   "EMP IDB_stations_me{1}_partNumbers{5}" : WString[40] = PLC "EMP IDB".stations.me[1].partNumbers[5], 1 s
   "EMP IDB_stations_me{1}_partNumbers{6}" : WString[40] = PLC "EMP IDB".stations.me[1].partNumbers[6], 1 s
   "EMP IDB_stations_me{1}_partNumbers{7}" : WString[40] = PLC "EMP IDB".stations.me[1].partNumbers[7], 1 s
   "EMP IDB_stations_me{2}_partNumbers{0}" : WString[40] = PLC "EMP IDB".stations.me[2].partNumbers[0], 1 s
   "EMP IDB_stations_me{2}_partNumbers{1}" : WString[40] = PLC "EMP IDB".stations.me[2].partNumbers[1], 1 s
   "EMP IDB_stations_me{2}_partNumbers{2}" : WString[40] = PLC "EMP IDB".stations.me[2].partNumbers[2], 1 s
   "EMP IDB_stations_me{2}_partNumbers{3}" : WString[40] = PLC "EMP IDB".stations.me[2].partNumbers[3], 1 s
   "EMP IDB_stations_me{2}_partNumbers{4}" : WString[40] = PLC "EMP IDB".stations.me[2].partNumbers[4], 1 s
   "EMP IDB_stations_me{2}_partNumbers{5}" : WString[40] = PLC "EMP IDB".stations.me[2].partNumbers[5], 1 s
   "EMP IDB_stations_me{2}_partNumbers{6}" : WString[40] = PLC "EMP IDB".stations.me[2].partNumbers[6], 1 s
   "EMP IDB_stations_me{2}_partNumbers{7}" : WString[40] = PLC "EMP IDB".stations.me[2].partNumbers[7], 1 s
   "EMP IDB_stations_me{3}_partOrdered{0}" : Bool = PLC "EMP IDB".stations.me[3].partOrdered[0], 1 s
   "EMP IDB_stations_me{3}_partOrdered{1}" : Bool = PLC "EMP IDB".stations.me[3].partOrdered[1], 1 s
   "EMP IDB_stations_me{3}_partOrdered{2}" : Bool = PLC "EMP IDB".stations.me[3].partOrdered[2], 1 s
   "EMP IDB_stations_me{3}_partOrdered{3}" : Bool = PLC "EMP IDB".stations.me[3].partOrdered[3], 1 s
   "EMP IDB_stations_me{3}_partOrdered{4}" : Bool = PLC "EMP IDB".stations.me[3].partOrdered[4], 1 s
   "EMP IDB_stations_me{3}_partOrdered{5}" : Bool = PLC "EMP IDB".stations.me[3].partOrdered[5], 1 s
   "EMP IDB_stations_me{3}_partOrdered{6}" : Bool = PLC "EMP IDB".stations.me[3].partOrdered[6], 1 s
   "EMP IDB_stations_me{3}_partOrdered{7}" : Bool = PLC "EMP IDB".stations.me[3].partOrdered[7], 1 s
   "EMP IDB_stations_me{4}_partNumbers{0}" : WString[40] = PLC "EMP IDB".stations.me[4].partNumbers[0], 1 s
   "EMP IDB_stations_me{4}_partNumbers{1}" : WString[40] = PLC "EMP IDB".stations.me[4].partNumbers[1], 1 s
   "EMP IDB_stations_me{4}_partNumbers{2}" : WString[40] = PLC "EMP IDB".stations.me[4].partNumbers[2], 1 s
   "EMP IDB_stations_me{4}_partNumbers{3}" : WString[40] = PLC "EMP IDB".stations.me[4].partNumbers[3], 1 s
   "EMP IDB_stations_me{4}_partNumbers{4}" : WString[40] = PLC "EMP IDB".stations.me[4].partNumbers[4], 1 s
   "EMP IDB_stations_me{4}_partNumbers{5}" : WString[40] = PLC "EMP IDB".stations.me[4].partNumbers[5], 1 s
   "EMP IDB_stations_me{4}_partNumbers{6}" : WString[40] = PLC "EMP IDB".stations.me[4].partNumbers[6], 1 s
   "EMP IDB_stations_me{4}_partNumbers{7}" : WString[40] = PLC "EMP IDB".stations.me[4].partNumbers[7], 1 s
   "EMP IDB_stations_me{5}_partNumbers{0}" : WString[40] = PLC "EMP IDB".stations.me[5].partNumbers[0], 1 s
   "EMP IDB_stations_me{5}_partNumbers{1}" : WString[40] = PLC "EMP IDB".stations.me[5].partNumbers[1], 1 s
   "EMP IDB_stations_me{5}_partNumbers{2}" : WString[40] = PLC "EMP IDB".stations.me[5].partNumbers[2], 1 s
   "EMP IDB_stations_me{5}_partNumbers{3}" : WString[40] = PLC "EMP IDB".stations.me[5].partNumbers[3], 1 s
   "EMP IDB_stations_me{5}_partNumbers{4}" : WString[40] = PLC "EMP IDB".stations.me[5].partNumbers[4], 1 s
   "EMP IDB_stations_me{5}_partNumbers{5}" : WString[40] = PLC "EMP IDB".stations.me[5].partNumbers[5], 1 s
   "EMP IDB_stations_me{5}_partNumbers{6}" : WString[40] = PLC "EMP IDB".stations.me[5].partNumbers[6], 1 s
   "EMP IDB_stations_me{5}_partNumbers{7}" : WString[40] = PLC "EMP IDB".stations.me[5].partNumbers[7], 1 s
   "EMP IDB_stations_me{6}_partNumbers{0}" : WString[40] = PLC "EMP IDB".stations.me[6].partNumbers[0], 1 s
   "EMP IDB_stations_me{6}_partNumbers{1}" : WString[40] = PLC "EMP IDB".stations.me[6].partNumbers[1], 1 s
   "EMP IDB_stations_me{6}_partNumbers{2}" : WString[40] = PLC "EMP IDB".stations.me[6].partNumbers[2], 1 s
   "EMP IDB_stations_me{6}_partNumbers{3}" : WString[40] = PLC "EMP IDB".stations.me[6].partNumbers[3], 1 s
   "EMP IDB_stations_me{6}_partNumbers{4}" : WString[40] = PLC "EMP IDB".stations.me[6].partNumbers[4], 1 s
   "EMP IDB_stations_me{6}_partNumbers{5}" : WString[40] = PLC "EMP IDB".stations.me[6].partNumbers[5], 1 s
   "EMP IDB_stations_me{6}_partNumbers{6}" : WString[40] = PLC "EMP IDB".stations.me[6].partNumbers[6], 1 s
   "EMP IDB_stations_me{6}_partNumbers{7}" : WString[40] = PLC "EMP IDB".stations.me[6].partNumbers[7], 1 s
   "EMP IDB_stations_me{7}_partNumbers{0}" : WString[40] = PLC "EMP IDB".stations.me[7].partNumbers[0], 1 s
   "EMP IDB_stations_me{7}_partNumbers{1}" : WString[40] = PLC "EMP IDB".stations.me[7].partNumbers[1], 1 s
   "EMP IDB_stations_me{7}_partNumbers{2}" : WString[40] = PLC "EMP IDB".stations.me[7].partNumbers[2], 1 s
   "EMP IDB_stations_me{7}_partNumbers{3}" : WString[40] = PLC "EMP IDB".stations.me[7].partNumbers[3], 1 s
   "EMP IDB_stations_me{7}_partNumbers{4}" : WString[40] = PLC "EMP IDB".stations.me[7].partNumbers[4], 1 s
   "EMP IDB_stations_me{7}_partNumbers{5}" : WString[40] = PLC "EMP IDB".stations.me[7].partNumbers[5], 1 s
   "EMP IDB_stations_me{7}_partNumbers{6}" : WString[40] = PLC "EMP IDB".stations.me[7].partNumbers[6], 1 s
   "EMP IDB_stations_me{7}_partNumbers{7}" : WString[40] = PLC "EMP IDB".stations.me[7].partNumbers[7], 1 s
   "EMP IDB_stations_me{8}_partNumbers{0}" : WString[40] = PLC "EMP IDB".stations.me[8].partNumbers[0], 1 s
   "EMP IDB_stations_me{8}_partNumbers{1}" : WString[40] = PLC "EMP IDB".stations.me[8].partNumbers[1], 1 s
   "EMP IDB_stations_me{8}_partNumbers{2}" : WString[40] = PLC "EMP IDB".stations.me[8].partNumbers[2], 1 s
   "EMP IDB_stations_me{8}_partNumbers{3}" : WString[40] = PLC "EMP IDB".stations.me[8].partNumbers[3], 1 s
   "EMP IDB_stations_me{8}_partNumbers{4}" : WString[40] = PLC "EMP IDB".stations.me[8].partNumbers[4], 1 s
   "EMP IDB_stations_me{8}_partNumbers{5}" : WString[40] = PLC "EMP IDB".stations.me[8].partNumbers[5], 1 s
   "EMP IDB_stations_me{8}_partNumbers{6}" : WString[40] = PLC "EMP IDB".stations.me[8].partNumbers[6], 1 s
   "EMP IDB_stations_me{8}_partNumbers{7}" : WString[40] = PLC "EMP IDB".stations.me[8].partNumbers[7], 1 s
   "EMP IDB_stations_me{9}_partNumbers{0}" : WString[40] = PLC "EMP IDB".stations.me[9].partNumbers[0], 1 s
   "EMP IDB_stations_me{9}_partNumbers{1}" : WString[40] = PLC "EMP IDB".stations.me[9].partNumbers[1], 1 s
   "EMP IDB_stations_me{9}_partNumbers{2}" : WString[40] = PLC "EMP IDB".stations.me[9].partNumbers[2], 1 s
   "EMP IDB_stations_me{9}_partNumbers{3}" : WString[40] = PLC "EMP IDB".stations.me[9].partNumbers[3], 1 s
   "EMP IDB_stations_me{9}_partNumbers{4}" : WString[40] = PLC "EMP IDB".stations.me[9].partNumbers[4], 1 s
   "EMP IDB_stations_me{9}_partNumbers{5}" : WString[40] = PLC "EMP IDB".stations.me[9].partNumbers[5], 1 s
   "EMP IDB_stations_me{9}_partNumbers{6}" : WString[40] = PLC "EMP IDB".stations.me[9].partNumbers[6], 1 s
   "EMP IDB_stations_me{9}_partNumbers{7}" : WString[40] = PLC "EMP IDB".stations.me[9].partNumbers[7], 1 s
   "EMP IDB_stations_me{10}_partNumbers{0}" : WString[40] = PLC "EMP IDB".stations.me[10].partNumbers[0], 1 s
   "EMP IDB_stations_me{10}_partNumbers{1}" : WString[40] = PLC "EMP IDB".stations.me[10].partNumbers[1], 1 s
   "EMP IDB_stations_me{10}_partNumbers{2}" : WString[40] = PLC "EMP IDB".stations.me[10].partNumbers[2], 1 s
   "EMP IDB_stations_me{10}_partNumbers{3}" : WString[40] = PLC "EMP IDB".stations.me[10].partNumbers[3], 1 s
   "EMP IDB_stations_me{10}_partNumbers{4}" : WString[40] = PLC "EMP IDB".stations.me[10].partNumbers[4], 1 s
   "EMP IDB_stations_me{10}_partNumbers{5}" : WString[40] = PLC "EMP IDB".stations.me[10].partNumbers[5], 1 s
   "EMP IDB_stations_me{10}_partNumbers{6}" : WString[40] = PLC "EMP IDB".stations.me[10].partNumbers[6], 1 s
   "EMP IDB_stations_me{10}_partNumbers{7}" : WString[40] = PLC "EMP IDB".stations.me[10].partNumbers[7], 1 s
   "EMP IDB_stations_me{11}_partNumbers{0}" : WString[40] = PLC "EMP IDB".stations.me[11].partNumbers[0], 1 s
   "EMP IDB_stations_me{11}_partNumbers{1}" : WString[40] = PLC "EMP IDB".stations.me[11].partNumbers[1], 1 s
   "EMP IDB_stations_me{11}_partNumbers{2}" : WString[40] = PLC "EMP IDB".stations.me[11].partNumbers[2], 1 s
   "EMP IDB_stations_me{11}_partNumbers{3}" : WString[40] = PLC "EMP IDB".stations.me[11].partNumbers[3], 1 s
   "EMP IDB_stations_me{11}_partNumbers{4}" : WString[40] = PLC "EMP IDB".stations.me[11].partNumbers[4], 1 s
   "EMP IDB_stations_me{11}_partNumbers{5}" : WString[40] = PLC "EMP IDB".stations.me[11].partNumbers[5], 1 s
   "EMP IDB_stations_me{11}_partNumbers{6}" : WString[40] = PLC "EMP IDB".stations.me[11].partNumbers[6], 1 s
   "EMP IDB_stations_me{11}_partNumbers{7}" : WString[40] = PLC "EMP IDB".stations.me[11].partNumbers[7], 1 s
   "EMP IDB_stations_me{12}_partNumbers{0}" : WString[40] = PLC "EMP IDB".stations.me[12].partNumbers[0], 1 s
   "EMP IDB_stations_me{12}_partNumbers{1}" : WString[40] = PLC "EMP IDB".stations.me[12].partNumbers[1], 1 s
   "EMP IDB_stations_me{12}_partNumbers{2}" : WString[40] = PLC "EMP IDB".stations.me[12].partNumbers[2], 1 s
   "EMP IDB_stations_me{12}_partNumbers{3}" : WString[40] = PLC "EMP IDB".stations.me[12].partNumbers[3], 1 s
   "EMP IDB_stations_me{12}_partNumbers{4}" : WString[40] = PLC "EMP IDB".stations.me[12].partNumbers[4], 1 s
   "EMP IDB_stations_me{12}_partNumbers{5}" : WString[40] = PLC "EMP IDB".stations.me[12].partNumbers[5], 1 s
   "EMP IDB_stations_me{12}_partNumbers{6}" : WString[40] = PLC "EMP IDB".stations.me[12].partNumbers[6], 1 s
   "EMP IDB_stations_me{12}_partNumbers{7}" : WString[40] = PLC "EMP IDB".stations.me[12].partNumbers[7], 1 s
   "EMP IDB_stations_me{13}_partNumbers{0}" : WString[40] = PLC "EMP IDB".stations.me[13].partNumbers[0], 1 s
   "EMP IDB_stations_me{13}_partNumbers{1}" : WString[40] = PLC "EMP IDB".stations.me[13].partNumbers[1], 1 s
   "EMP IDB_stations_me{13}_partNumbers{2}" : WString[40] = PLC "EMP IDB".stations.me[13].partNumbers[2], 1 s
   "EMP IDB_stations_me{13}_partNumbers{3}" : WString[40] = PLC "EMP IDB".stations.me[13].partNumbers[3], 1 s
   "EMP IDB_stations_me{13}_partNumbers{4}" : WString[40] = PLC "EMP IDB".stations.me[13].partNumbers[4], 1 s
   "EMP IDB_stations_me{13}_partNumbers{5}" : WString[40] = PLC "EMP IDB".stations.me[13].partNumbers[5], 1 s
   "EMP IDB_stations_me{13}_partNumbers{6}" : WString[40] = PLC "EMP IDB".stations.me[13].partNumbers[6], 1 s
   "EMP IDB_stations_me{13}_partNumbers{7}" : WString[40] = PLC "EMP IDB".stations.me[13].partNumbers[7], 1 s
   "EMP IDB_stations_me{14}_partNumbers{0}" : WString[40] = PLC "EMP IDB".stations.me[14].partNumbers[0], 1 s
   "EMP IDB_stations_me{14}_partNumbers{1}" : WString[40] = PLC "EMP IDB".stations.me[14].partNumbers[1], 1 s
   "EMP IDB_stations_me{14}_partNumbers{2}" : WString[40] = PLC "EMP IDB".stations.me[14].partNumbers[2], 1 s
   "EMP IDB_stations_me{14}_partNumbers{3}" : WString[40] = PLC "EMP IDB".stations.me[14].partNumbers[3], 1 s
   "EMP IDB_stations_me{14}_partNumbers{4}" : WString[40] = PLC "EMP IDB".stations.me[14].partNumbers[4], 1 s
   "EMP IDB_stations_me{14}_partNumbers{5}" : WString[40] = PLC "EMP IDB".stations.me[14].partNumbers[5], 1 s
   "EMP IDB_stations_me{14}_partNumbers{6}" : WString[40] = PLC "EMP IDB".stations.me[14].partNumbers[6], 1 s
   "EMP IDB_stations_me{14}_partNumbers{7}" : WString[40] = PLC "EMP IDB".stations.me[14].partNumbers[7], 1 s
   "EMP IDB_stations_me{15}_partNumbers{0}" : WString[40] = PLC "EMP IDB".stations.me[15].partNumbers[0], 1 s
   "EMP IDB_stations_me{15}_partNumbers{1}" : WString[40] = PLC "EMP IDB".stations.me[15].partNumbers[1], 1 s
   "EMP IDB_stations_me{15}_partNumbers{2}" : WString[40] = PLC "EMP IDB".stations.me[15].partNumbers[2], 1 s
   "EMP IDB_stations_me{15}_partNumbers{3}" : WString[40] = PLC "EMP IDB".stations.me[15].partNumbers[3], 1 s
   "EMP IDB_stations_me{15}_partNumbers{4}" : WString[40] = PLC "EMP IDB".stations.me[15].partNumbers[4], 1 s
   "EMP IDB_stations_me{15}_partNumbers{5}" : WString[40] = PLC "EMP IDB".stations.me[15].partNumbers[5], 1 s
   "EMP IDB_stations_me{15}_partNumbers{6}" : WString[40] = PLC "EMP IDB".stations.me[15].partNumbers[6], 1 s
   "EMP IDB_stations_me{15}_partNumbers{7}" : WString[40] = PLC "EMP IDB".stations.me[15].partNumbers[7], 1 s
   "EMP IDB_stations_me{16}_partNumbers{0}" : WString[40] = PLC "EMP IDB".stations.me[16].partNumbers[0], 1 s
   "EMP IDB_stations_me{16}_partNumbers{1}" : WString[40] = PLC "EMP IDB".stations.me[16].partNumbers[1], 1 s
   "EMP IDB_stations_me{16}_partNumbers{2}" : WString[40] = PLC "EMP IDB".stations.me[16].partNumbers[2], 1 s
   "EMP IDB_stations_me{16}_partNumbers{3}" : WString[40] = PLC "EMP IDB".stations.me[16].partNumbers[3], 1 s
   "EMP IDB_stations_me{16}_partNumbers{4}" : WString[40] = PLC "EMP IDB".stations.me[16].partNumbers[4], 1 s
   "EMP IDB_stations_me{16}_partNumbers{5}" : WString[40] = PLC "EMP IDB".stations.me[16].partNumbers[5], 1 s
   "EMP IDB_stations_me{16}_partNumbers{6}" : WString[40] = PLC "EMP IDB".stations.me[16].partNumbers[6], 1 s
   "EMP IDB_stations_me{16}_partNumbers{7}" : WString[40] = PLC "EMP IDB".stations.me[16].partNumbers[7], 1 s
   "EMP IDB_stations_me{17}_partNumbers{0}" : WString[40] = PLC "EMP IDB".stations.me[17].partNumbers[0], 1 s
   "EMP IDB_stations_me{17}_partNumbers{1}" : WString[40] = PLC "EMP IDB".stations.me[17].partNumbers[1], 1 s
   "EMP IDB_stations_me{17}_partNumbers{2}" : WString[40] = PLC "EMP IDB".stations.me[17].partNumbers[2], 1 s
   "EMP IDB_stations_me{17}_partNumbers{3}" : WString[40] = PLC "EMP IDB".stations.me[17].partNumbers[3], 1 s
   "EMP IDB_stations_me{17}_partNumbers{4}" : WString[40] = PLC "EMP IDB".stations.me[17].partNumbers[4], 1 s
   "EMP IDB_stations_me{17}_partNumbers{5}" : WString[40] = PLC "EMP IDB".stations.me[17].partNumbers[5], 1 s
   "EMP IDB_stations_me{17}_partNumbers{6}" : WString[40] = PLC "EMP IDB".stations.me[17].partNumbers[6], 1 s
   "EMP IDB_stations_me{17}_partNumbers{7}" : WString[40] = PLC "EMP IDB".stations.me[17].partNumbers[7], 1 s
   "EMP IDB_stations_me{18}_partNumbers{0}" : WString[40] = PLC "EMP IDB".stations.me[18].partNumbers[0], 1 s
   "EMP IDB_stations_me{18}_partNumbers{1}" : WString[40] = PLC "EMP IDB".stations.me[18].partNumbers[1], 1 s
   "EMP IDB_stations_me{18}_partNumbers{2}" : WString[40] = PLC "EMP IDB".stations.me[18].partNumbers[2], 1 s
   "EMP IDB_stations_me{18}_partNumbers{3}" : WString[40] = PLC "EMP IDB".stations.me[18].partNumbers[3], 1 s
   "EMP IDB_stations_me{18}_partNumbers{4}" : WString[40] = PLC "EMP IDB".stations.me[18].partNumbers[4], 1 s
   "EMP IDB_stations_me{18}_partNumbers{5}" : WString[40] = PLC "EMP IDB".stations.me[18].partNumbers[5], 1 s
   "EMP IDB_stations_me{18}_partNumbers{6}" : WString[40] = PLC "EMP IDB".stations.me[18].partNumbers[6], 1 s
   "EMP IDB_stations_me{18}_partNumbers{7}" : WString[40] = PLC "EMP IDB".stations.me[18].partNumbers[7], 1 s
   "EMP IDB_stations_me{19}_partNumbers{0}" : WString[40] = PLC "EMP IDB".stations.me[19].partNumbers[0], 1 s
   "EMP IDB_stations_me{19}_partNumbers{1}" : WString[40] = PLC "EMP IDB".stations.me[19].partNumbers[1], 1 s
   "EMP IDB_stations_me{19}_partNumbers{2}" : WString[40] = PLC "EMP IDB".stations.me[19].partNumbers[2], 1 s
   "EMP IDB_stations_me{19}_partNumbers{3}" : WString[40] = PLC "EMP IDB".stations.me[19].partNumbers[3], 1 s
   "EMP IDB_stations_me{19}_partNumbers{4}" : WString[40] = PLC "EMP IDB".stations.me[19].partNumbers[4], 1 s
   "EMP IDB_stations_me{19}_partNumbers{5}" : WString[40] = PLC "EMP IDB".stations.me[19].partNumbers[5], 1 s
   "EMP IDB_stations_me{19}_partNumbers{6}" : WString[40] = PLC "EMP IDB".stations.me[19].partNumbers[6], 1 s
   "EMP IDB_stations_me{19}_partNumbers{7}" : WString[40] = PLC "EMP IDB".stations.me[19].partNumbers[7], 1 s
   "EMP IDB_stations_me{20}_partNumbers{0}" : WString[40] = PLC "EMP IDB".stations.me[20].partNumbers[0], 1 s
   "EMP IDB_stations_me{20}_partNumbers{1}" : WString[40] = PLC "EMP IDB".stations.me[20].partNumbers[1], 1 s
   "EMP IDB_stations_me{20}_partNumbers{2}" : WString[40] = PLC "EMP IDB".stations.me[20].partNumbers[2], 1 s
   "EMP IDB_stations_me{20}_partNumbers{3}" : WString[40] = PLC "EMP IDB".stations.me[20].partNumbers[3], 1 s
   "EMP IDB_stations_me{20}_partNumbers{4}" : WString[40] = PLC "EMP IDB".stations.me[20].partNumbers[4], 1 s
   "EMP IDB_stations_me{20}_partNumbers{5}" : WString[40] = PLC "EMP IDB".stations.me[20].partNumbers[5], 1 s
   "EMP IDB_stations_me{20}_partNumbers{6}" : WString[40] = PLC "EMP IDB".stations.me[20].partNumbers[6], 1 s
   "EMP IDB_stations_me{20}_partNumbers{7}" : WString[40] = PLC "EMP IDB".stations.me[20].partNumbers[7], 1 s
   "EMP IDB_stations_me{21}_partNumbers{0}" : WString[40] = PLC "EMP IDB".stations.me[21].partNumbers[0], 1 s
   "EMP IDB_stations_me{21}_partNumbers{1}" : WString[40] = PLC "EMP IDB".stations.me[21].partNumbers[1], 1 s
   "EMP IDB_stations_me{21}_partNumbers{2}" : WString[40] = PLC "EMP IDB".stations.me[21].partNumbers[2], 1 s
   "EMP IDB_stations_me{21}_partNumbers{3}" : WString[40] = PLC "EMP IDB".stations.me[21].partNumbers[3], 1 s
   "EMP IDB_stations_me{21}_partNumbers{4}" : WString[40] = PLC "EMP IDB".stations.me[21].partNumbers[4], 1 s
   "EMP IDB_stations_me{21}_partNumbers{5}" : WString[40] = PLC "EMP IDB".stations.me[21].partNumbers[5], 1 s
   "EMP IDB_stations_me{21}_partNumbers{6}" : WString[40] = PLC "EMP IDB".stations.me[21].partNumbers[6], 1 s
   "EMP IDB_stations_me{21}_partNumbers{7}" : WString[40] = PLC "EMP IDB".stations.me[21].partNumbers[7], 1 s
   "EMP IDB_stations_me{22}_partNumbers{0}" : WString[40] = PLC "EMP IDB".stations.me[22].partNumbers[0], 1 s
   "EMP IDB_stations_me{22}_partNumbers{1}" : WString[40] = PLC "EMP IDB".stations.me[22].partNumbers[1], 1 s
   "EMP IDB_stations_me{22}_partNumbers{2}" : WString[40] = PLC "EMP IDB".stations.me[22].partNumbers[2], 1 s
   "EMP IDB_stations_me{22}_partNumbers{3}" : WString[40] = PLC "EMP IDB".stations.me[22].partNumbers[3], 1 s
   "EMP IDB_stations_me{22}_partNumbers{4}" : WString[40] = PLC "EMP IDB".stations.me[22].partNumbers[4], 1 s
   "EMP IDB_stations_me{22}_partNumbers{5}" : WString[40] = PLC "EMP IDB".stations.me[22].partNumbers[5], 1 s
   "EMP IDB_stations_me{22}_partNumbers{6}" : WString[40] = PLC "EMP IDB".stations.me[22].partNumbers[6], 1 s
   "EMP IDB_stations_me{22}_partNumbers{7}" : WString[40] = PLC "EMP IDB".stations.me[22].partNumbers[7], 1 s
   "EMP IDB_stations_me{23}_partNumbers{0}" : WString[40] = PLC "EMP IDB".stations.me[23].partNumbers[0], 1 s
   "EMP IDB_stations_me{23}_partNumbers{1}" : WString[40] = PLC "EMP IDB".stations.me[23].partNumbers[1], 1 s
   "EMP IDB_stations_me{23}_partNumbers{2}" : WString[40] = PLC "EMP IDB".stations.me[23].partNumbers[2], 1 s
   "EMP IDB_stations_me{23}_partNumbers{3}" : WString[40] = PLC "EMP IDB".stations.me[23].partNumbers[3], 1 s
   "EMP IDB_stations_me{23}_partNumbers{4}" : WString[40] = PLC "EMP IDB".stations.me[23].partNumbers[4], 1 s
   "EMP IDB_stations_me{23}_partNumbers{5}" : WString[40] = PLC "EMP IDB".stations.me[23].partNumbers[5], 1 s
   "EMP IDB_stations_me{23}_partNumbers{6}" : WString[40] = PLC "EMP IDB".stations.me[23].partNumbers[6], 1 s
   "EMP IDB_stations_me{23}_partNumbers{7}" : WString[40] = PLC "EMP IDB".stations.me[23].partNumbers[7], 1 s
   "EMP IDB_stations_me{3}_partNumbers{0}" : WString[40] = PLC "EMP IDB".stations.me[3].partNumbers[0], 1 s
   "EMP IDB_stations_me{3}_partNumbers{1}" : WString[40] = PLC "EMP IDB".stations.me[3].partNumbers[1], 1 s
   "EMP IDB_stations_me{3}_partNumbers{2}" : WString[40] = PLC "EMP IDB".stations.me[3].partNumbers[2], 1 s
   "EMP IDB_stations_me{3}_partNumbers{3}" : WString[40] = PLC "EMP IDB".stations.me[3].partNumbers[3], 1 s
   "EMP IDB_stations_me{3}_partNumbers{4}" : WString[40] = PLC "EMP IDB".stations.me[3].partNumbers[4], 1 s
   "EMP IDB_stations_me{3}_partNumbers{5}" : WString[40] = PLC "EMP IDB".stations.me[3].partNumbers[5], 1 s
   "EMP IDB_stations_me{3}_partNumbers{6}" : WString[40] = PLC "EMP IDB".stations.me[3].partNumbers[6], 1 s
   "EMP IDB_stations_me{3}_partNumbers{7}" : WString[40] = PLC "EMP IDB".stations.me[3].partNumbers[7], 1 s

text list "Station Selection Single": 0 'Select a Station to View'; 1 'Assignments'

recipe "VOLVO 16 01": Button 0 <- "EMP IDB_stations_me{0}_partNumbers{0}", Button 1 <- "EMP IDB_stations_me{0}_partNumbers{1}", Button 2 <- "EMP IDB_stations_me{0}_partNumbers{2}", Button 3 <- "EMP IDB_stations_me{0}_partNumbers{3}", Button 4 <- "EMP IDB_stations_me{0}_partNumbers{4}", Button 5 <- "EMP IDB_stations_me{0}_partNumbers{5}", Button 6 <- "EMP IDB_stations_me{0}_partNumbers{6}", Button 7 <- "EMP IDB_stations_me{0}_partNumbers{7}"

recipe "VOLVO 16 02": Button 0 <- "EMP IDB_stations_me{1}_partNumbers{0}", Button 1 <- "EMP IDB_stations_me{1}_partNumbers{1}", Button 2 <- "EMP IDB_stations_me{1}_partNumbers{2}", Button 3 <- "EMP IDB_stations_me{1}_partNumbers{3}", Button 4 <- "EMP IDB_stations_me{1}_partNumbers{4}", Button 5 <- "EMP IDB_stations_me{1}_partNumbers{5}", Button 6 <- "EMP IDB_stations_me{1}_partNumbers{6}", Button 7 <- "EMP IDB_stations_me{1}_partNumbers{7}"

recipe "VOLVO 16 03": Button 0 <- "EMP IDB_stations_me{2}_partNumbers{0}", Button 1 <- "EMP IDB_stations_me{2}_partNumbers{1}", Button 2 <- "EMP IDB_stations_me{2}_partNumbers{2}", Button 3 <- "EMP IDB_stations_me{2}_partNumbers{3}", Button 4 <- "EMP IDB_stations_me{2}_partNumbers{4}", Button 5 <- "EMP IDB_stations_me{2}_partNumbers{5}", Button 6 <- "EMP IDB_stations_me{2}_partNumbers{6}", Button 7 <- "EMP IDB_stations_me{2}_partNumbers{7}"

recipe "VOLVO 16 04": Button 0 <- "EMP IDB_stations_me{3}_partNumbers{0}", Button 1 <- "EMP IDB_stations_me{3}_partNumbers{1}", Button 2 <- "EMP IDB_stations_me{3}_partNumbers{2}", Button 3 <- "EMP IDB_stations_me{3}_partNumbers{3}", Button 4 <- "EMP IDB_stations_me{3}_partNumbers{4}", Button 5 <- "EMP IDB_stations_me{3}_partNumbers{5}", Button 6 <- "EMP IDB_stations_me{3}_partNumbers{6}", Button 7 <- "EMP IDB_stations_me{3}_partNumbers{7}"

recipe "VOLVO 16 05": Button 0 <- "EMP IDB_stations_me{4}_partNumbers{0}", Button 1 <- "EMP IDB_stations_me{4}_partNumbers{1}", Button 2 <- "EMP IDB_stations_me{4}_partNumbers{2}", Button 3 <- "EMP IDB_stations_me{4}_partNumbers{3}", Button 4 <- "EMP IDB_stations_me{4}_partNumbers{4}", Button 5 <- "EMP IDB_stations_me{4}_partNumbers{5}", Button 6 <- "EMP IDB_stations_me{4}_partNumbers{6}", Button 7 <- "EMP IDB_stations_me{4}_partNumbers{7}"

recipe "VOLVO 16 06": Button 0 <- "EMP IDB_stations_me{5}_partNumbers{0}", Button 1 <- "EMP IDB_stations_me{5}_partNumbers{1}", Button 2 <- "EMP IDB_stations_me{5}_partNumbers{2}", Button 3 <- "EMP IDB_stations_me{5}_partNumbers{3}", Button 4 <- "EMP IDB_stations_me{5}_partNumbers{4}", Button 5 <- "EMP IDB_stations_me{5}_partNumbers{5}", Button 6 <- "EMP IDB_stations_me{5}_partNumbers{6}", Button 7 <- "EMP IDB_stations_me{5}_partNumbers{7}"

recipe "VOLVO 16 07": Button 0 <- "EMP IDB_stations_me{6}_partNumbers{0}", Button 1 <- "EMP IDB_stations_me{6}_partNumbers{1}", Button 2 <- "EMP IDB_stations_me{6}_partNumbers{2}", Button 3 <- "EMP IDB_stations_me{6}_partNumbers{3}", Button 4 <- "EMP IDB_stations_me{6}_partNumbers{4}", Button 5 <- "EMP IDB_stations_me{6}_partNumbers{5}", Button 6 <- "EMP IDB_stations_me{6}_partNumbers{6}", Button 7 <- "EMP IDB_stations_me{6}_partNumbers{7}"

recipe "VOLVO 16 08": Button 0 <- "EMP IDB_stations_me{7}_partNumbers{0}", Button 1 <- "EMP IDB_stations_me{7}_partNumbers{1}", Button 2 <- "EMP IDB_stations_me{7}_partNumbers{2}", Button 3 <- "EMP IDB_stations_me{7}_partNumbers{3}", Button 4 <- "EMP IDB_stations_me{7}_partNumbers{4}", Button 5 <- "EMP IDB_stations_me{7}_partNumbers{5}", Button 6 <- "EMP IDB_stations_me{7}_partNumbers{6}", Button 7 <- "EMP IDB_stations_me{7}_partNumbers{7}"

recipe "VOLVO 16 09": Button 0 <- "EMP IDB_stations_me{8}_partNumbers{0}", Button 1 <- "EMP IDB_stations_me{8}_partNumbers{1}", Button 2 <- "EMP IDB_stations_me{8}_partNumbers{2}", Button 3 <- "EMP IDB_stations_me{8}_partNumbers{3}", Button 4 <- "EMP IDB_stations_me{8}_partNumbers{4}", Button 5 <- "EMP IDB_stations_me{8}_partNumbers{5}", Button 6 <- "EMP IDB_stations_me{8}_partNumbers{6}", Button 7 <- "EMP IDB_stations_me{8}_partNumbers{7}"

recipe "VOLVO 16 10": Button 0 <- "EMP IDB_stations_me{9}_partNumbers{0}", Button 1 <- "EMP IDB_stations_me{9}_partNumbers{1}", Button 2 <- "EMP IDB_stations_me{9}_partNumbers{2}", Button 3 <- "EMP IDB_stations_me{9}_partNumbers{3}", Button 4 <- "EMP IDB_stations_me{9}_partNumbers{4}", Button 5 <- "EMP IDB_stations_me{9}_partNumbers{5}", Button 6 <- "EMP IDB_stations_me{9}_partNumbers{6}", Button 7 <- "EMP IDB_stations_me{9}_partNumbers{7}"

recipe "VOLVO 16 11": Button 0 <- "EMP IDB_stations_me{10}_partNumbers{0}", Button 1 <- "EMP IDB_stations_me{10}_partNumbers{1}", Button 2 <- "EMP IDB_stations_me{10}_partNumbers{2}", Button 3 <- "EMP IDB_stations_me{10}_partNumbers{3}", Button 4 <- "EMP IDB_stations_me{10}_partNumbers{4}", Button 5 <- "EMP IDB_stations_me{10}_partNumbers{5}", Button 6 <- "EMP IDB_stations_me{10}_partNumbers{6}", Button 7 <- "EMP IDB_stations_me{10}_partNumbers{7}"

recipe "CHM 01": Button 0 <- "EMP IDB_stations_me{11}_partNumbers{0}", Button 1 <- "EMP IDB_stations_me{11}_partNumbers{1}", Button 2 <- "EMP IDB_stations_me{11}_partNumbers{2}", Button 3 <- "EMP IDB_stations_me{11}_partNumbers{3}", Button 4 <- "EMP IDB_stations_me{11}_partNumbers{4}", Button 5 <- "EMP IDB_stations_me{11}_partNumbers{5}", Button 6 <- "EMP IDB_stations_me{11}_partNumbers{6}", Button 7 <- "EMP IDB_stations_me{11}_partNumbers{7}"

recipe "CHM 02": Button 0 <- "EMP IDB_stations_me{12}_partNumbers{0}", Button 1 <- "EMP IDB_stations_me{12}_partNumbers{1}", Button 2 <- "EMP IDB_stations_me{12}_partNumbers{2}", Button 3 <- "EMP IDB_stations_me{12}_partNumbers{3}", Button 4 <- "EMP IDB_stations_me{12}_partNumbers{4}", Button 5 <- "EMP IDB_stations_me{12}_partNumbers{5}", Button 6 <- "EMP IDB_stations_me{12}_partNumbers{6}", Button 7 <- "EMP IDB_stations_me{12}_partNumbers{7}"

recipe "CHM 03": Button 0 <- "EMP IDB_stations_me{13}_partNumbers{0}", Button 1 <- "EMP IDB_stations_me{13}_partNumbers{1}", Button 2 <- "EMP IDB_stations_me{13}_partNumbers{2}", Button 3 <- "EMP IDB_stations_me{13}_partNumbers{3}", Button 4 <- "EMP IDB_stations_me{13}_partNumbers{4}", Button 5 <- "EMP IDB_stations_me{13}_partNumbers{5}", Button 6 <- "EMP IDB_stations_me{13}_partNumbers{6}", Button 7 <- "EMP IDB_stations_me{13}_partNumbers{7}"

recipe "CHM 04": Button 0 <- "EMP IDB_stations_me{14}_partNumbers{0}", Button 1 <- "EMP IDB_stations_me{14}_partNumbers{1}", Button 2 <- "EMP IDB_stations_me{14}_partNumbers{2}", Button 3 <- "EMP IDB_stations_me{14}_partNumbers{3}", Button 4 <- "EMP IDB_stations_me{14}_partNumbers{4}", Button 5 <- "EMP IDB_stations_me{14}_partNumbers{5}", Button 6 <- "EMP IDB_stations_me{14}_partNumbers{6}", Button 7 <- "EMP IDB_stations_me{14}_partNumbers{7}"

recipe "CHM 05": Button 0 <- "EMP IDB_stations_me{15}_partNumbers{0}", Button 1 <- "EMP IDB_stations_me{15}_partNumbers{1}", Button 2 <- "EMP IDB_stations_me{15}_partNumbers{2}", Button 3 <- "EMP IDB_stations_me{15}_partNumbers{3}", Button 4 <- "EMP IDB_stations_me{15}_partNumbers{4}", Button 5 <- "EMP IDB_stations_me{15}_partNumbers{5}", Button 6 <- "EMP IDB_stations_me{15}_partNumbers{6}", Button 7 <- "EMP IDB_stations_me{15}_partNumbers{7}"

recipe "CDO 01": Button 0 <- "EMP IDB_stations_me{16}_partNumbers{0}", Button 1 <- "EMP IDB_stations_me{16}_partNumbers{1}", Button 2 <- "EMP IDB_stations_me{16}_partNumbers{2}", Button 3 <- "EMP IDB_stations_me{16}_partNumbers{3}", Button 4 <- "EMP IDB_stations_me{16}_partNumbers{4}", Button 5 <- "EMP IDB_stations_me{16}_partNumbers{5}", Button 6 <- "EMP IDB_stations_me{16}_partNumbers{6}", Button 7 <- "EMP IDB_stations_me{16}_partNumbers{7}"

recipe "CDO 02": Button 0 <- "EMP IDB_stations_me{17}_partNumbers{0}", Button 1 <- "EMP IDB_stations_me{17}_partNumbers{1}", Button 2 <- "EMP IDB_stations_me{17}_partNumbers{2}", Button 3 <- "EMP IDB_stations_me{17}_partNumbers{3}", Button 4 <- "EMP IDB_stations_me{17}_partNumbers{4}", Button 5 <- "EMP IDB_stations_me{17}_partNumbers{5}", Button 6 <- "EMP IDB_stations_me{17}_partNumbers{6}", Button 7 <- "EMP IDB_stations_me{17}_partNumbers{7}"

recipe "CDO 03": Button 0 <- "EMP IDB_stations_me{18}_partNumbers{0}", Button 1 <- "EMP IDB_stations_me{18}_partNumbers{1}", Button 2 <- "EMP IDB_stations_me{18}_partNumbers{2}", Button 3 <- "EMP IDB_stations_me{18}_partNumbers{3}", Button 4 <- "EMP IDB_stations_me{18}_partNumbers{4}", Button 5 <- "EMP IDB_stations_me{18}_partNumbers{5}", Button 6 <- "EMP IDB_stations_me{18}_partNumbers{6}", Button 7 <- "EMP IDB_stations_me{18}_partNumbers{7}"

recipe "BFL 01": Button 0 <- "EMP IDB_stations_me{19}_partNumbers{0}", Button 1 <- "EMP IDB_stations_me{19}_partNumbers{1}", Button 2 <- "EMP IDB_stations_me{19}_partNumbers{2}", Button 3 <- "EMP IDB_stations_me{19}_partNumbers{3}", Button 4 <- "EMP IDB_stations_me{19}_partNumbers{4}", Button 5 <- "EMP IDB_stations_me{19}_partNumbers{5}", Button 6 <- "EMP IDB_stations_me{19}_partNumbers{6}", Button 7 <- "EMP IDB_stations_me{19}_partNumbers{7}"

recipe "BFL 02": Button 0 <- "EMP IDB_stations_me{20}_partNumbers{0}", Button 1 <- "EMP IDB_stations_me{20}_partNumbers{1}", Button 2 <- "EMP IDB_stations_me{20}_partNumbers{2}", Button 3 <- "EMP IDB_stations_me{20}_partNumbers{3}", Button 4 <- "EMP IDB_stations_me{20}_partNumbers{4}", Button 5 <- "EMP IDB_stations_me{20}_partNumbers{5}", Button 6 <- "EMP IDB_stations_me{20}_partNumbers{6}", Button 7 <- "EMP IDB_stations_me{20}_partNumbers{7}"

recipe "BFL 03": Button 0 <- "EMP IDB_stations_me{21}_partNumbers{0}", Button 1 <- "EMP IDB_stations_me{21}_partNumbers{1}", Button 2 <- "EMP IDB_stations_me{21}_partNumbers{2}", Button 3 <- "EMP IDB_stations_me{21}_partNumbers{3}", Button 4 <- "EMP IDB_stations_me{21}_partNumbers{4}", Button 5 <- "EMP IDB_stations_me{21}_partNumbers{5}", Button 6 <- "EMP IDB_stations_me{21}_partNumbers{6}", Button 7 <- "EMP IDB_stations_me{21}_partNumbers{7}"

recipe "LGS 01": Button 0 <- "EMP IDB_stations_me{22}_partNumbers{0}", Button 1 <- "EMP IDB_stations_me{22}_partNumbers{1}", Button 2 <- "EMP IDB_stations_me{22}_partNumbers{2}", Button 3 <- "EMP IDB_stations_me{22}_partNumbers{3}", Button 4 <- "EMP IDB_stations_me{22}_partNumbers{4}", Button 5 <- "EMP IDB_stations_me{22}_partNumbers{5}", Button 6 <- "EMP IDB_stations_me{22}_partNumbers{6}", Button 7 <- "EMP IDB_stations_me{22}_partNumbers{7}"

recipe "LGS 02": Button 0 <- "EMP IDB_stations_me{23}_partNumbers{0}", Button 1 <- "EMP IDB_stations_me{23}_partNumbers{1}", Button 2 <- "EMP IDB_stations_me{23}_partNumbers{2}", Button 3 <- "EMP IDB_stations_me{23}_partNumbers{3}", Button 4 <- "EMP IDB_stations_me{23}_partNumbers{4}", Button 5 <- "EMP IDB_stations_me{23}_partNumbers{5}", Button 6 <- "EMP IDB_stations_me{23}_partNumbers{6}", Button 7 <- "EMP IDB_stations_me{23}_partNumbers{7}"

screen "1 PART CALL" 1366x768
   on GenerateScreen: SetTag("HMI_screenNumber", 1)
   Rectangle "Settings Tab Background" at 682,0 size 684x68
      Appearance <- "HMI_screenNumber"
   Rectangle "Part Call Tab Background" at 0,0 size 685x68
      Appearance <- "HMI_screenNumber"
   Rectangle "Settings Tab Border Hide" at 685,61 size 678x20
      Visibility <- "HMI_screenNumber"
   Rectangle "Part Call Tab Border Hide" at 3,61 size 679x20
      Visibility <- "HMI_screenNumber"
   Button "Settings Screen" at 683,0 size 683x68; TextOff 'SETTINGS'; Authorization "User administration"
      on Release: ActivateScreen("2 SETTINGS", 0)
   Button "Part Call Screen" at 0,0 size 683x68; TextOff 'PART CALL'
      on Release: ActivateScreen("1 PART CALL", 0)
   TextField "Header Line" at 32,112 size 216x53; Text 'LINE'
   TextField "Header Drop Zone" at 238,112 size 236x53; Text 'DROP ZONE'
   TextField "Header Part Number" at 474,112 size 648x53; Text 'PART NUMBER'
   TextField "Header Time" at 1112,112 size 222x53; Text 'TIME'
   ScreenModuleView "TableRow00" at 27,170 size 1312x52; ScreenModuleType ""
      Guid_{11997190-27688} <- "HMI_partCall_row{0}"
      on Guid_{11997190-83214}: ActivateScreen("3 BARCODE", 0)
   ScreenModuleView "TableRow01" at 27,222 size 1312x52; ScreenModuleType ""
      Guid_{11997190-27688} <- "HMI_partCall_row{1}"
      on Guid_{11997190-83214}: ActivateScreen("3 BARCODE", 0)
   ScreenModuleView "TableRow02" at 27,274 size 1312x52; ScreenModuleType ""
      Guid_{11997190-27688} <- "HMI_partCall_row{2}"
      on Guid_{11997190-83214}: ActivateScreen("3 BARCODE", 0)
   ScreenModuleView "TableRow03" at 27,326 size 1312x52; ScreenModuleType ""
      Guid_{11997190-27688} <- "HMI_partCall_row{3}"
      on Guid_{11997190-83214}: ActivateScreen("3 BARCODE", 0)
   ScreenModuleView "TableRow04" at 27,378 size 1312x52; ScreenModuleType ""
      Guid_{11997190-27688} <- "HMI_partCall_row{4}"
      on Guid_{11997190-83214}: ActivateScreen("3 BARCODE", 0)
   ScreenModuleView "TableRow05" at 27,430 size 1312x52; ScreenModuleType ""
      Guid_{11997190-27688} <- "HMI_partCall_row{5}"
      on Guid_{11997190-83214}: ActivateScreen("3 BARCODE", 0)
   ScreenModuleView "TableRow06" at 27,482 size 1312x52; ScreenModuleType ""
      Guid_{11997190-27688} <- "HMI_partCall_row{6}"
      on Guid_{11997190-83214}: ActivateScreen("3 BARCODE", 0)
   ScreenModuleView "TableRow07" at 27,534 size 1312x52; ScreenModuleType ""
      Guid_{11997190-27688} <- "HMI_partCall_row{7}"
      on Guid_{11997190-83214}: ActivateScreen("3 BARCODE", 0)
   ScreenModuleView "TableRow08" at 27,586 size 1312x52; ScreenModuleType ""
      Guid_{11997190-27688} <- "HMI_partCall_row{8}"
      on Guid_{11997190-83214}: ActivateScreen("3 BARCODE", 0)
   ScreenModuleView "TableRow09" at 27,638 size 1312x52; ScreenModuleType ""
      Guid_{11997190-27688} <- "HMI_partCall_row{9}"
      on Guid_{11997190-83214}: ActivateScreen("3 BARCODE", 0)
   ScreenModuleView "TableRow10" at 27,690 size 1312x52; ScreenModuleType ""
      Guid_{11997190-27688} <- "HMI_partCall_row{10}"
      on Guid_{11997190-83214}: ActivateScreen("3 BARCODE", 0)

screen "2 SETTINGS" 1366x768
   on GenerateScreen: SetTag("HMI_screenNumber", 2)
   Rectangle "Part Call Nave Panel" at 0,0 size 455x68
      Appearance <- "HMI_screenNumber"
   Rectangle "Settings Nav Panel" at 452,0 size 462x68
      Appearance <- "HMI_screenNumber"
   Rectangle "Network Health Nav Panel" at 911,0 size 455x68
      Appearance <- "HMI_screenNumber"
   Rectangle "Part Call Border Hide" at 3,60 size 449x20
      Visibility <- "HMI_screenNumber"
   Rectangle "Settings Border Hide" at 455,60 size 456x20
      Visibility <- "HMI_screenNumber"
   Rectangle "Network Health Border Hide" at 914,60 size 449x20
      Visibility <- "HMI_screenNumber"
   Button "Part Call Screen" at 0,0 size 455x68; TextOff 'PART CALL'
      on Release: ActivateScreen("1 PART CALL", 0)
   Button "Settings Screen" at 455,0 size 460x68; TextOff 'SETTINGS'
      on Release: ActivateScreen("2 SETTINGS", 0)
   Button "Network Health Screen" at 914,0 size 452x68; TextOff 'NW HEALTH'
      on Release: ActivateScreen("4 NETWORK HEALTH", 0)
   Rectangle "Station Assignment Table BG Full" at 793,120 size 533x630
      Visibility <- "HMI_settings_stations_selCount"
   TextField "Current Station Single" at 803,130 size 513x45; Text 'Text'
      Visibility <- "HMI_settings_stations_selCount"
   TextField "Hide Line and Drop Zone Multi" at 803,181 size 513x40; Text 'select single station for Line and Drop Zone'
      Visibility <- "HMI_settings_stations_selCount"
   GraphicView "KP8 Image" at 496,327 size 275x412; Picture "kp8 image"
   Rectangle "Station Assignment Table BG Mini" at 793,120 size 533x65
      Visibility <- "HMI_settings_stations_selCount"
   ScreenModuleView "PB: Set PN" at 50,130 size 414x45; Guid_{11997190-63616} 'Assign Part Number'; ScreenModuleType ""
      Guid_{11997190-63605} <- "HMI_settings_partNumber_assign"
   ScreenModuleView "PN IO Field" at 50,180 size 414x50; ScreenModuleType ""
      Guid_{11997190-63113} <- "HMI_settings_partNumber_ioField"
   ScreenModuleView "PB: Set Allotted" at 494,130 size 137x45; Guid_{11997190-63616} 'Allotted'; ScreenModuleType ""
      Guid_{11997190-63605} <- "HMI_settings_alotted_assign"
   ScreenModuleView "PB: Set Critical" at 636,130 size 137x45; Guid_{11997190-63616} 'Crititcal'; ScreenModuleType ""
      Guid_{11997190-63605} <- "HMI_settings_critical_assign"
   ScreenModuleView "Alotted Time IO Field" at 494,180 size 137x50; ScreenModuleType ""
      Guid_{11997190-63269} <- "HMI_settings_alotted_ioField"
   ScreenModuleView "Critical Time IO Field" at 636,180 size 137x50; ScreenModuleType ""
      Guid_{11997190-63269} <- "HMI_settings_critical_ioField"
   ScreenModuleView "PB: Select KP8 Buttons" at 493,270 size 284x45; Guid_{11997190-63616} 'Select Buttons'; ScreenModuleType ""
      Guid_{11997190-63605} <- "HMI_settings_kp8_selectButtons"
   ScreenModuleView "KP8 00: RESET" at 641,614 size 68x66; ScreenModuleType ""
      Guid_{11997190-57808} <- "HMI_settings_kp8_buttons{0}"
   ScreenModuleView "KP8 01" at 641,535 size 68x66; ScreenModuleType ""
      Guid_{11997190-57808} <- "HMI_settings_kp8_buttons{1}"
   ScreenModuleView "KP8 02" at 641,459 size 68x66; ScreenModuleType ""
      Guid_{11997190-57808} <- "HMI_settings_kp8_buttons{2}"
   ScreenModuleView "KP8 03" at 641,383 size 68x66; ScreenModuleType ""
      Guid_{11997190-57808} <- "HMI_settings_kp8_buttons{3}"
   ScreenModuleView "KP8 04: STOP RUNTIME" at 557,614 size 68x66; ScreenModuleType ""
      on Guid_{11997190-59171}: StopRuntime(0)
      Guid_{11997190-57808} <- "HMI_settings_kp8_buttons{4}"
   ScreenModuleView "KP8 05" at 557,535 size 68x66; ScreenModuleType ""
      Guid_{11997190-57808} <- "HMI_settings_kp8_buttons{5}"
   ScreenModuleView "KP8 06" at 557,459 size 68x66; ScreenModuleType ""
      Guid_{11997190-57808} <- "HMI_settings_kp8_buttons{6}"
   ScreenModuleView "KP8 07" at 557,383 size 68x66; ScreenModuleType ""
      Guid_{11997190-57808} <- "HMI_settings_kp8_buttons{7}"
   ScreenModuleView "PB: Previous Group" at 50,270 size 65x45; Guid_{11997190-63799} "Up"; ScreenModuleType ""
      Guid_{11997190-63779} <- "HMI_settings_stations_prevGroup"
   ScreenModuleView "PB: Select All Stations" at 120,270 size 274x45; Guid_{11997190-63616} 'Select Stations'; ScreenModuleType ""
      Guid_{11997190-63605} <- "HMI_settings_stations_selectAll"
   ScreenModuleView "PB: Next Group" at 399,270 size 65x45; Guid_{11997190-63799} "Down"; ScreenModuleType ""
      Guid_{11997190-63779} <- "HMI_settings_stations_nextGroup"
   ScreenModuleView "Station 00 Select" at 50,320 size 205x65; ScreenModuleType ""
      Guid_{11997190-57808} <- "HMI_settings_stations_selectBtns{0}"
   ScreenModuleView "Station 01 Select" at 260,320 size 205x65; ScreenModuleType ""
      Guid_{11997190-57808} <- "HMI_settings_stations_selectBtns{1}"
   ScreenModuleView "Station 02 Select" at 50,391 size 205x65; ScreenModuleType ""
      Guid_{11997190-57808} <- "HMI_settings_stations_selectBtns{2}"
   ScreenModuleView "Station 03 Select" at 260,391 size 205x65; ScreenModuleType ""
      Guid_{11997190-57808} <- "HMI_settings_stations_selectBtns{3}"
   ScreenModuleView "Station 04 Select" at 50,462 size 205x65; ScreenModuleType ""
      Guid_{11997190-57808} <- "HMI_settings_stations_selectBtns{4}"
   ScreenModuleView "Station 05 Select" at 260,462 size 205x65; ScreenModuleType ""
      Guid_{11997190-57808} <- "HMI_settings_stations_selectBtns{5}"
   ScreenModuleView "Station 06 Select" at 50,533 size 205x65; ScreenModuleType ""
      Guid_{11997190-57808} <- "HMI_settings_stations_selectBtns{6}"
   ScreenModuleView "Station 07 Select" at 260,533 size 205x65; ScreenModuleType ""
      Guid_{11997190-57808} <- "HMI_settings_stations_selectBtns{7}"
   ScreenModuleView "Station 08 Select" at 50,604 size 205x65; ScreenModuleType ""
      Guid_{11997190-57808} <- "HMI_settings_stations_selectBtns{8}"
   ScreenModuleView "Station 09 Select" at 260,604 size 205x65; ScreenModuleType ""
      Guid_{11997190-57808} <- "HMI_settings_stations_selectBtns{9}"
   ScreenModuleView "Station 10 Select" at 50,675 size 205x65; ScreenModuleType ""
      Guid_{11997190-57808} <- "HMI_settings_stations_selectBtns{10}"
   ScreenModuleView "Station 11 Select" at 260,675 size 205x65; ScreenModuleType ""
      Guid_{11997190-57808} <- "HMI_settings_stations_selectBtns{11}"
   ScreenModuleView "Line Label" at 803,181 size 267x40; ScreenModuleType ""
      Guid_{11997190-64598} <- "HMI_settings_viewingStation_lineData"
   ScreenModuleView "Drop Zone Label" at 1076,181 size 240x40; ScreenModuleType ""
      Guid_{11997190-64802} <- "HMI_settings_viewingStation_dzData"
   ScreenModuleView "PB: Previous Station" at 803,130 size 65x45; Guid_{11997190-63799} "Left"; ScreenModuleType ""
      Guid_{11997190-63779} <- "HMI_settings_viewingStation_previous"
   TextField "Current Station Multi" at 873,130 size 373x45; Text 'Assignments'
      Visibility <- "HMI_settings_stations_selCount"
   ScreenModuleView "PB: Next Station" at 1251,130 size 65x45; Guid_{11997190-63799} "Right"; ScreenModuleType ""
      Guid_{11997190-63779} <- "HMI_settings_viewingStation_next"
   TextField "Button Column Header" at 803,226 size 75x40; Text 'Btn'
      Visibility <- "HMI_settings_stations_selCount"
   TextField "Timer Column Header" at 872,226 size 128x40; Text 'Times'
      Visibility <- "HMI_settings_stations_selCount"
   TextField "Part Number Column Header" at 993,226 size 323x40; Text 'Part Number'
      Visibility <- "HMI_settings_stations_selCount"
   ScreenModuleView "Button 00 Details" at 803,271 size 513x74; ScreenModuleType ""
      Guid_{11997190-60358} <- "HMI_settings_viewingStation_btns{0}"
   ScreenModuleView "Button 01 Details" at 803,350 size 513x74; ScreenModuleType ""
      Guid_{11997190-60358} <- "HMI_settings_viewingStation_btns{1}"
   ScreenModuleView "Button 02 Details" at 803,429 size 513x74; ScreenModuleType ""
      Guid_{11997190-60358} <- "HMI_settings_viewingStation_btns{2}"
   ScreenModuleView "Button 03 Details" at 803,508 size 513x74; ScreenModuleType ""
      Guid_{11997190-60358} <- "HMI_settings_viewingStation_btns{3}"
   ScreenModuleView "Button 04 Details" at 803,587 size 513x74; ScreenModuleType ""
      Guid_{11997190-60358} <- "HMI_settings_viewingStation_btns{4}"
   ScreenModuleView "Button 05 Details" at 803,666 size 513x74; ScreenModuleType ""
      Guid_{11997190-60358} <- "HMI_settings_viewingStation_btns{5}"

SlideinScreen "GraphX_Slidein_Bottom" 1366x80
   ScreenModuleView "Top" at 0,0 size 227x80; Guid_{11997190-63799} "Top"; ScreenModuleType ""
      Guid_{11997190-63779} <- "HMI_tableNav_top"
   ScreenModuleView "Page Up" at 227,0 size 228x80; Guid_{11997190-63799} "pageUp"; ScreenModuleType ""
      Guid_{11997190-63779} <- "HMI_tableNav_pageUp"
   ScreenModuleView "Line Up" at 455,0 size 228x80; Guid_{11997190-63799} "Up"; ScreenModuleType ""
      Guid_{11997190-63779} <- "HMI_tableNav_lineUp"
   ScreenModuleView "Line Down" at 683,0 size 228x80; Guid_{11997190-63799} "Down"; ScreenModuleType ""
      Guid_{11997190-63779} <- "HMI_tableNav_lineDown"
   ScreenModuleView "Page Down" at 911,0 size 228x80; Guid_{11997190-63799} "PageDown"; ScreenModuleType ""
      Guid_{11997190-63779} <- "HMI_tableNav_pageDown"
   ScreenModuleView "Bottom" at 1138,0 size 228x80; Guid_{11997190-63799} "Bottom"; ScreenModuleType ""
      Guid_{11997190-63779} <- "HMI_tableNav_bottom"
   TextField "Text field_1" at 0,0 size 1366x80; Text 'NOT USED'
      Visibility <- "HMI_screenNumber"

SlideinScreen "GraphX_Slidein_Right" 449x768
   ScreenModuleView "Station Sim_1" at 5,5 size 106x232; ScreenModuleType ""
      Guid_{11997190-89108} <- "HMI_simStations_stations{0}"
   ScreenModuleView "Station Sim_2" at 116,5 size 106x232; ScreenModuleType ""
      Guid_{11997190-89108} <- "HMI_simStations_me{1}"
   ScreenModuleView "Station Sim_3" at 227,5 size 106x232; ScreenModuleType ""
      Guid_{11997190-89108} <- "HMI_simStations_me{2}"
   ScreenModuleView "Station Sim_4" at 338,5 size 106x232; ScreenModuleType ""
      Guid_{11997190-89108} <- "HMI_simStations_me{3}"
   ScreenModuleView "Station Sim_5" at 5,242 size 106x232; ScreenModuleType ""
      Guid_{11997190-89108} <- "HMI_simStations_me{4}"
   ScreenModuleView "Station Sim_6" at 5,479 size 106x232; ScreenModuleType ""
      Guid_{11997190-89108} <- "HMI_simStations_me{8}"
   ScreenModuleView "Station Sim_7" at 116,242 size 106x232; ScreenModuleType ""
      Guid_{11997190-89108} <- "HMI_simStations_me{5}"
   ScreenModuleView "Station Sim_8" at 227,242 size 106x232; ScreenModuleType ""
      Guid_{11997190-89108} <- "HMI_simStations_me{6}"
   ScreenModuleView "Station Sim_9" at 338,242 size 106x232; ScreenModuleType ""
      Guid_{11997190-89108} <- "HMI_simStations_me{7}"
   ScreenModuleView "Station Sim_10" at 116,479 size 106x232; ScreenModuleType ""
      Guid_{11997190-89108} <- "HMI_simStations_me{9}"
   ScreenModuleView "Station Sim_11" at 227,478 size 106x232; ScreenModuleType ""
      Guid_{11997190-89108} <- "HMI_simStations_me{10}"
   ScreenModuleView "Station Sim_12" at 338,477 size 106x232; ScreenModuleType ""
      Guid_{11997190-89108} <- "HMI_simStations_me{11}"
   ScreenModuleView "PB: Graphic/Text List_1" at 5,716 size 65x45; Guid_{11997190-63799} "Up"; ScreenModuleType ""
      Guid_{11997190-63779} <- "HMI_simStations_up"
   ScreenModuleView "PB: Graphic/Text List_2" at 379,716 size 65x45; Guid_{11997190-63799} "Down"; ScreenModuleType ""
      Guid_{11997190-63779} <- "HMI_simStations_down"

screen "3 BARCODE" 1366x768
   on GenerateScreen: SetTag("HMI_screenNumber", 3)
   Rectangle "Nav Panel 02" at 682,700 size 684x68
      Appearance <- "HMI_screenNumber"
   Rectangle "Nav Panel 01" at 0,700 size 685x68
      Appearance <- "HMI_screenNumber"
   Rectangle "Nav Panel 03 Top Border Hide" at 685,700 size 678x3
      Visibility <- "HMI_screenNumber"
   Rectangle "Nav Panel 01 Top Border Hide" at 3,700 size 679x3
      Visibility <- "HMI_screenNumber"
   Button "Settings Screen" at 683,700 size 683x68; TextOff 'SETTINGS'; Authorization "User administration"
      on Release: ActivateScreen("2 SETTINGS", 0)
   Button "Part Call Screen" at 0,700 size 683x68; TextOff 'PART CALL'
      on Release: ActivateScreen("1 PART CALL", 0)
   Button "btCancel" at 685,431 size 649x68; TextOff 'CANCEL'
      on Release: ActivateScreen("1 PART CALL", 0)
   Button "btPartOrdered" at 32,431 size 648x68; TextOff 'ORDERED'
      on Release: SetBit("ordered"); ActivateScreen("1 PART CALL", 0)
   TextField "tfBarcodeDisplay" at 32,220 size 1302x206; Text 'Text'
   TextField "tfPartNumberDisplay" at 32,160 size 1302x53; Text 'BARCODE FOR PART NUMBER'

